// TIA Portal project "Inteligenta_szklarnia" (V15.1) (continued)
REGION Network 2: Warunki dla których okna są otwierane
   // Gdy uruchomiony jest tryb automatyczny, wartość CO2 w szklarni powinna się mieścić w zakresie nastawionego stężenia CO2 +- wartość histerezy. Okna są otwierane po spełnieniu następujących warunków: 1) gdy użytkownik załączył tryb okien na HMI, 2) gdy stężenie CO2 jest poza tym wymaganym przedziałem, 3) gdy stężenie CO2 poza szklarnią jest większe, jeśli chcemy zwiększyć ilość CO2 w szklarni oraz mniejsze, jeśli chcemy zmniejszyć ilość CO2 w szklarni, 4) gdy temperatura poza szklarnią mieści się w przedziale +-5°C temperatury nastawionej, 5) gdy wiatr wieje z prędkością nie większą niż 35km/h. Jeśli stężenie CO2 wzrośnie do niebezpiecznego poziomu 975ppm, okna również są otwierane bez względu na warunki zewnętrzne. W trybie manualnym okna otwierane są od razu po naciśnięciu przycisku do niego przypisanego.
   RUNG wire#powerrail
      Contact( #czy_automatyczny )
      I_Contact( #czy_manualny )
      wire#w1
      Contact( "HMI".System_okien_auto )
      { S7_Templates := "SrcType := Int" } LE_Contact(in1 := "Wejscia_PLC".Czujnik_wiatru, in2 := 35)
      wire#w2
      { S7_Templates := "SrcType := Int" } LT_Contact(in1 := #Histereza_plus, in2 := "HMI".Poziom_CO2_auto)
      { S7_Templates := "SrcType := Int" } GT_Contact(in1 := "Wejscia_PLC".Wewnetrzny_czujnik_CO2, in2 := "Wejscia_PLC".Zewnetrzny_czujnik_CO2)
      wire#w3
      { S7_Templates := "SrcType := Real" } InRange(min := #Zakres_temp_dol, in := "Wejscia_PLC".Temperatura_zewnetrzna, max := #Zakres_temp_gora)
      wire#w4
      I_Contact( "Siłownik_okien_zamykanie" )
      Coil( "Siłownik_okien_otwieranie" )
   END_RUNG
   RUNG wire#w2
      { S7_Templates := "SrcType := Int" } GT_Contact(in1 := #Histereza_minus, in2 := "Wejscia_PLC".Wewnetrzny_czujnik_CO2)
      { S7_Templates := "SrcType := Int" } LT_Contact(in1 := "Wejscia_PLC".Wewnetrzny_czujnik_CO2, in2 := "Wejscia_PLC".Zewnetrzny_czujnik_CO2)
   END_RUNG wire#w3
   RUNG wire#w1
      { S7_Templates := "SrcType := Int" } GE_Contact(in1 := "Wejscia_PLC".Wewnetrzny_czujnik_CO2, in2 := 975)
      { S7_Templates := "SrcType := Int" } GT_Contact(in1 := "Wejscia_PLC".Wewnetrzny_czujnik_CO2, in2 := "Wejscia_PLC".Zewnetrzny_czujnik_CO2)
   END_RUNG wire#w4
   RUNG wire#powerrail
      Contact( #czy_manualny )
      I_Contact( #czy_automatyczny )
      Contact( "HMI".Otwarcie_okien_manual )
   END_RUNG wire#w4
   // the same network as SCL:
   "Siłownik_okien_otwieranie" := ((#czy_automatyczny AND NOT #czy_manualny AND (("HMI".System_okien_auto AND ("Wejscia_PLC".Czujnik_wiatru <= 35) AND (((#Histereza_plus < "HMI".Poziom_CO2_auto) AND ("Wejscia_PLC".Wewnetrzny_czujnik_CO2 > "Wejscia_PLC".Zewnetrzny_czujnik_CO2)) OR ((#Histereza_minus > "Wejscia_PLC".Wewnetrzny_czujnik_CO2) AND ("Wejscia_PLC".Wewnetrzny_czujnik_CO2 < "Wejscia_PLC".Zewnetrzny_czujnik_CO2))) AND (#Zakres_temp_dol <= "Wejscia_PLC".Temperatura_zewnetrzna) AND ("Wejscia_PLC".Temperatura_zewnetrzna <= #Zakres_temp_gora)) OR (("Wejscia_PLC".Wewnetrzny_czujnik_CO2 >= 975) AND ("Wejscia_PLC".Wewnetrzny_czujnik_CO2 > "Wejscia_PLC".Zewnetrzny_czujnik_CO2)))) OR (#czy_manualny AND NOT #czy_automatyczny AND "HMI".Otwarcie_okien_manual)) AND NOT "Siłownik_okien_zamykanie";
END_REGION

REGION Network 3: Warunki dla których okna są zamykane
   // W trybie automatycznym okna są zamykane: 1) gdy tryb okien został wyłączony przez użytkownika, 2) gdy stężenie CO2 w szklarni wynosi zadaną wartość tego parametru +- histereza, 3) gdy stężenie CO2 poza szklarnią jest mniejsze, niż wewnątrz, jeśli chcemy zwiększyć jego ilość oraz większe, gdy chcemy zmniejszyć jego ilość, 4) gdy tempperatura zewnętrzna różni się o ponad 5°C od zadanej, 5) gdy wiatr wieje z prędkością większą niż 35km/h, 6) gdy stężenie CO2 w szklarni nie przekracza 955ppm lub przekracza, ale stężenie CO2 poza szklarnią jest większe. W trybie manualnym okna są zamykane, gdy przełączk na HMI znajdzie się w pozycji "ZAMKNIĘTE".
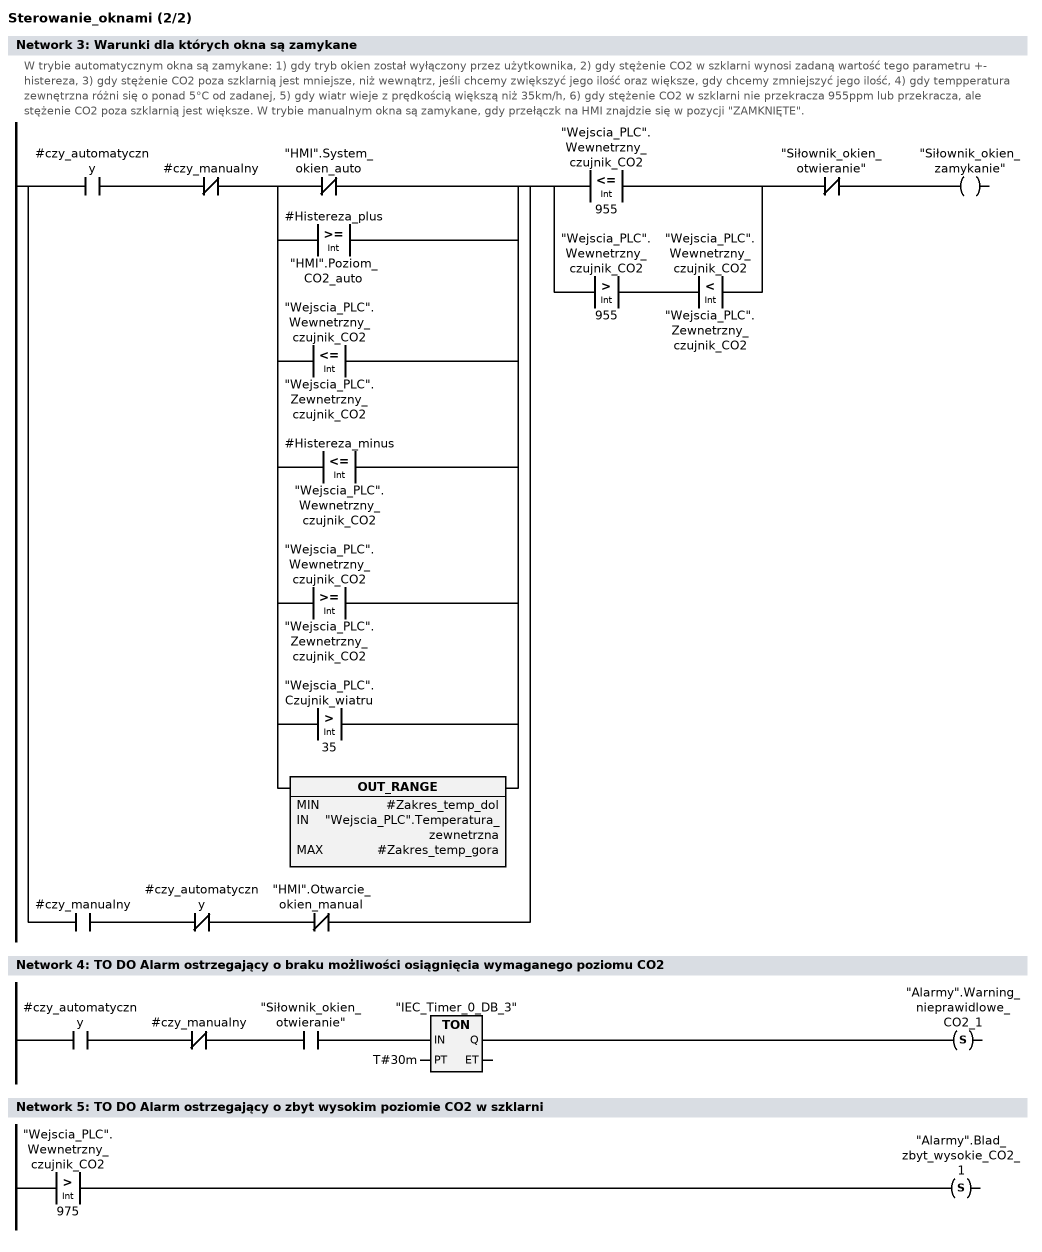
   "Siłownik_okien_zamykanie" := ((#czy_automatyczny AND NOT #czy_manualny AND (NOT "HMI".System_okien_auto OR (#Histereza_plus >= "HMI".Poziom_CO2_auto) OR ("Wejscia_PLC".Wewnetrzny_czujnik_CO2 <= "Wejscia_PLC".Zewnetrzny_czujnik_CO2) OR (#Histereza_minus <= "Wejscia_PLC".Wewnetrzny_czujnik_CO2) OR ("Wejscia_PLC".Wewnetrzny_czujnik_CO2 >= "Wejscia_PLC".Zewnetrzny_czujnik_CO2) OR ("Wejscia_PLC".Czujnik_wiatru > 35) OR ("Wejscia_PLC".Temperatura_zewnetrzna < #Zakres_temp_dol) OR ("Wejscia_PLC".Temperatura_zewnetrzna > #Zakres_temp_gora))) OR (#czy_manualny AND NOT #czy_automatyczny AND NOT "HMI".Otwarcie_okien_manual)) AND (("Wejscia_PLC".Wewnetrzny_czujnik_CO2 <= 955) OR (("Wejscia_PLC".Wewnetrzny_czujnik_CO2 > 955) AND ("Wejscia_PLC".Wewnetrzny_czujnik_CO2 < "Wejscia_PLC".Zewnetrzny_czujnik_CO2))) AND NOT "Siłownik_okien_otwieranie";
END_REGION

REGION Network 4: TO DO Alarm ostrzegający o braku możliwości osiągnięcia wymaganego poziomu CO2
   "IEC_Timer_0_DB_3".TON(IN := #czy_automatyczny AND NOT #czy_manualny AND "Siłownik_okien_otwieranie",
                          PT := T#30m);
   IF "IEC_Timer_0_DB_3".Q THEN "Alarmy".Warning_nieprawidlowe_CO2_1 := TRUE; END_IF;
END_REGION

REGION Network 5: TO DO Alarm ostrzegający o zbyt wysokim poziomie CO2 w szklarni
   RUNG wire#powerrail
      { S7_Templates := "SrcType := Int" } GT_Contact(in1 := "Wejscia_PLC".Wewnetrzny_czujnik_CO2, in2 := 975)
      S_Coil( "Alarmy".Blad_zbyt_wysokie_CO2_1 )
   END_RUNG
   // the same network as SCL:
   IF "Wejscia_PLC".Wewnetrzny_czujnik_CO2 > 975 THEN "Alarmy".Blad_zbyt_wysokie_CO2_1 := TRUE; END_IF;
END_REGION
END_FUNCTION

FUNCTION "SYMULACJA" : Void   // FC9, LAD
{ S7_Optimized_Access := 'TRUE' }
VERSION : 0.1
   VAR_INPUT
      counters : Bool;
   END_VAR
   VAR_TEMP
      temperatura_temp : Real;
      roznica_temperatur : Real;
      "wilgotność powietrza_temp" : Int;
      wilgotnosc_gleby_temp : Int;
      stezenie_CO2 : Int;
      natezenie_swiatla_temp : Int;
      odsloniecie_okna_temp : Real;
      pedkosc_wiatru_temp : Real;
      rand : Real;
      error : Bool;
      status : Int;
      sub_status : Int;
      rolety_temp : Real;
      test1 : Real;
   END_VAR
   VAR_TEMP   // added for the SCL form of the ladder/FBD networks
      _w1 : Bool;
   END_VAR
BEGIN

REGION Network 1: blok oblicza roznice temperatur
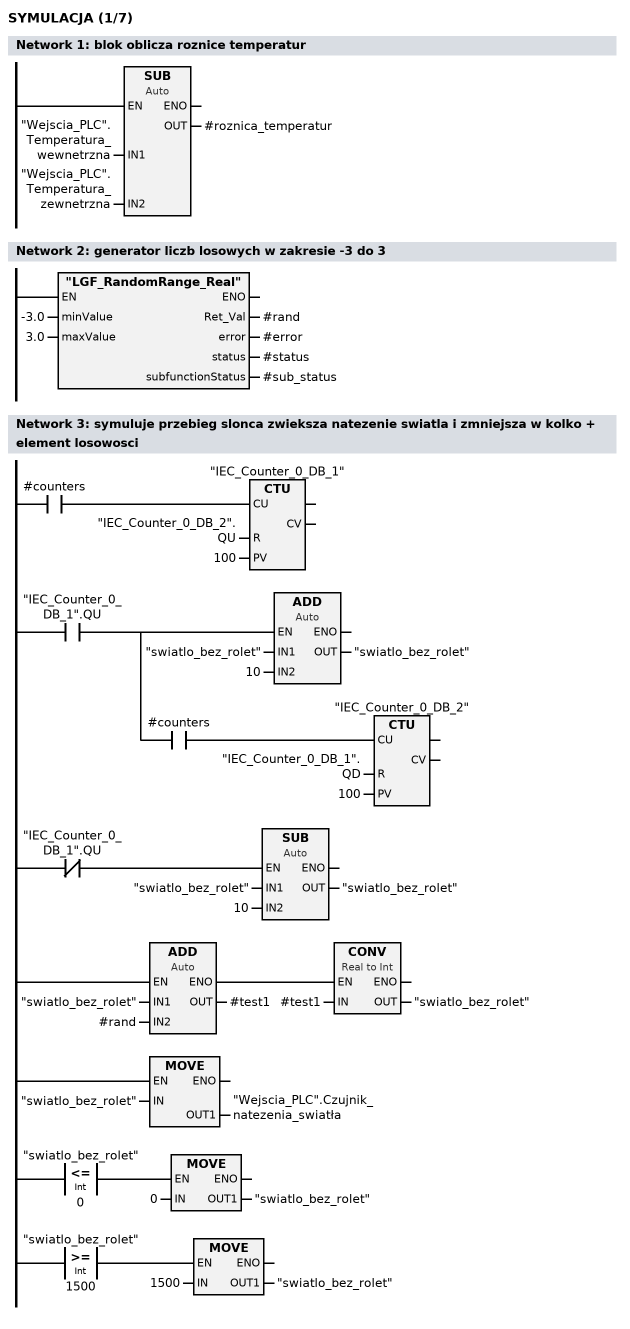
   RUNG wire#powerrail
      { S7_GenerateENO := "TRUE" } Sub(in1 := "Wejscia_PLC".Temperatura_wewnetrzna, in2 := "Wejscia_PLC".Temperatura_zewnetrzna, out => #roznica_temperatur)
   END_RUNG
   // the same network as SCL:
   #roznica_temperatur := "Wejscia_PLC".Temperatura_wewnetrzna - "Wejscia_PLC".Temperatura_zewnetrzna;
END_REGION

REGION Network 2: generator liczb losowych w zakresie -3 do 3
   RUNG wire#powerrail
      "LGF_RandomRange_Real"(minValue := -3.0, maxValue := 3.0, Ret_Val => #rand, error => #error, status => #status, subfunctionStatus => #sub_status)
   END_RUNG
   // the same network as SCL:
   #rand := "LGF_RandomRange_Real"(minValue := -3.0,
                           maxValue := 3.0,
                           error => #error,
                           status => #status,
                           subfunctionStatus => #sub_status);
END_REGION

REGION Network 3: symuluje przebieg slonca zwieksza natezenie swiatla i zmniejsza w kolko + element losowosci
   // ENO of a box is taken as its EN; it also drops when the box reports an error
   "IEC_Counter_0_DB_1".CTU(CU := #counters, R := "IEC_Counter_0_DB_2".QU, PV := 100);
   IF "IEC_Counter_0_DB_1".QU THEN "swiatlo_bez_rolet" := "swiatlo_bez_rolet" + 10; END_IF;
   "IEC_Counter_0_DB_2".CTU(CU := "IEC_Counter_0_DB_1".QU AND #counters,
                           R := "IEC_Counter_0_DB_1".QD,
                           PV := 100);
   IF NOT "IEC_Counter_0_DB_1".QU THEN "swiatlo_bez_rolet" := "swiatlo_bez_rolet" - 10; END_IF;
   #test1 := "swiatlo_bez_rolet" + #rand;
   "swiatlo_bez_rolet" := REAL_TO_INT(#test1);
   "Wejscia_PLC".Czujnik_natezenia_swiatła := "swiatlo_bez_rolet";
   IF "swiatlo_bez_rolet" <= 0 THEN "swiatlo_bez_rolet" := 0; END_IF;
   IF "swiatlo_bez_rolet" >= 1500 THEN "swiatlo_bez_rolet" := 1500; END_IF;
END_REGION

REGION Network 4: funkcja oblicza liniową zależność natężenia światła od zasłonięcia rolet
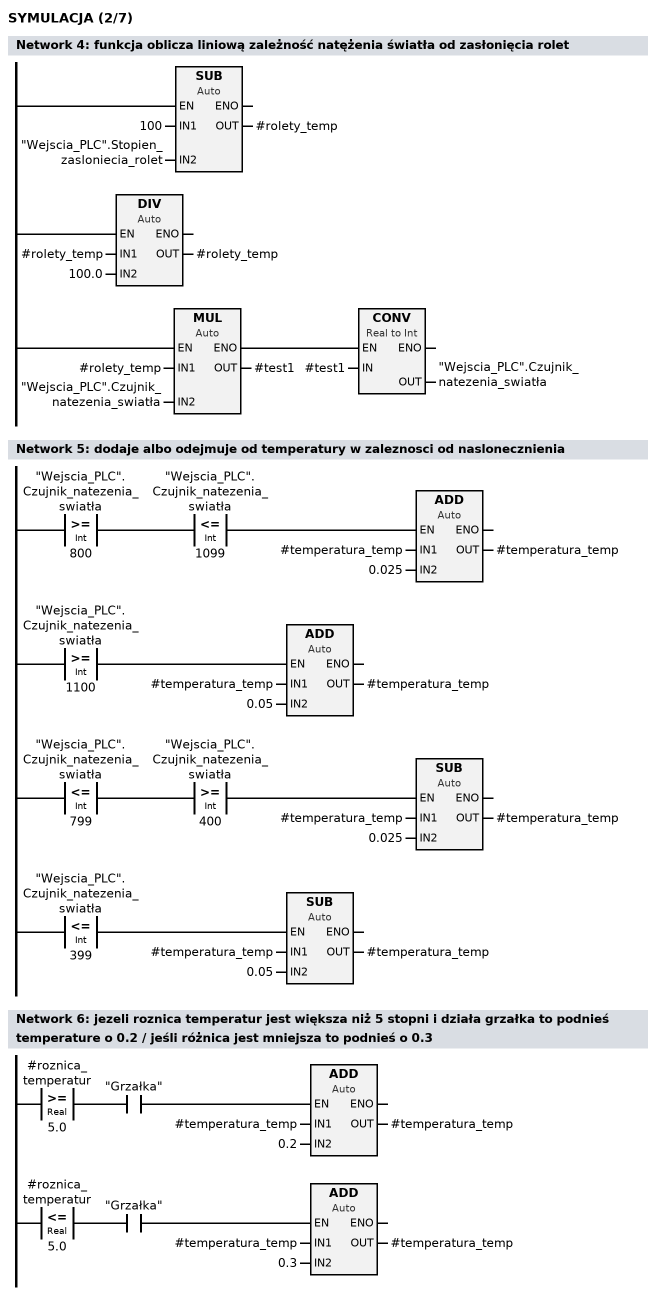
   RUNG wire#powerrail
      { S7_GenerateENO := "TRUE" } Sub(in1 := 100, in2 := "Wejscia_PLC".Stopien_zasloniecia_rolet, out => #rolety_temp)
   END_RUNG
   RUNG wire#powerrail
      { S7_GenerateENO := "TRUE" } Div(in1 := #rolety_temp, in2 := 100.0, out => #rolety_temp)
   END_RUNG
   RUNG wire#powerrail
      { S7_GenerateENO := "TRUE" } Mul(in1 := #rolety_temp, in2 := "Wejscia_PLC".Czujnik_natezenia_swiatła, out => #test1)
      { S7_Templates := "[SrcType := Real, DestType := Int]"; S7_GenerateENO := "TRUE" } Convert(in := #test1, out => "Wejscia_PLC".Czujnik_natezenia_swiatła)
   END_RUNG
   // the same network as SCL:
   // ENO of a box is taken as its EN; it also drops when the box reports an error
   #rolety_temp := 100 - "Wejscia_PLC".Stopien_zasloniecia_rolet;
   #rolety_temp := #rolety_temp / 100.0;
   #test1 := #rolety_temp * "Wejscia_PLC".Czujnik_natezenia_swiatła;
   "Wejscia_PLC".Czujnik_natezenia_swiatła := REAL_TO_INT(#test1);
END_REGION

REGION Network 5: dodaje albo odejmuje od temperatury w zaleznosci od naslonecznienia
   RUNG wire#powerrail
      { S7_Templates := "SrcType := Int" } GE_Contact(in1 := "Wejscia_PLC".Czujnik_natezenia_swiatła, in2 := 800)
      { S7_Templates := "SrcType := Int" } LE_Contact(in1 := "Wejscia_PLC".Czujnik_natezenia_swiatła, in2 := 1099)
      { S7_GenerateENO := "TRUE" } Add(in1 := #temperatura_temp, in2 := 0.025, out => #temperatura_temp)
   END_RUNG
   RUNG wire#powerrail
      { S7_Templates := "SrcType := Int" } GE_Contact(in1 := "Wejscia_PLC".Czujnik_natezenia_swiatła, in2 := 1100)
      { S7_GenerateENO := "TRUE" } Add(in1 := #temperatura_temp, in2 := 0.05, out => #temperatura_temp)
   END_RUNG
   RUNG wire#powerrail
      { S7_Templates := "SrcType := Int" } LE_Contact(in1 := "Wejscia_PLC".Czujnik_natezenia_swiatła, in2 := 799)
      { S7_Templates := "SrcType := Int" } GE_Contact(in1 := "Wejscia_PLC".Czujnik_natezenia_swiatła, in2 := 400)
      { S7_GenerateENO := "TRUE" } Sub(in1 := #temperatura_temp, in2 := 0.025, out => #temperatura_temp)
   END_RUNG
   RUNG wire#powerrail
      { S7_Templates := "SrcType := Int" } LE_Contact(in1 := "Wejscia_PLC".Czujnik_natezenia_swiatła, in2 := 399)
      { S7_GenerateENO := "TRUE" } Sub(in1 := #temperatura_temp, in2 := 0.05, out => #temperatura_temp)
   END_RUNG
   // the same network as SCL:
   IF ("Wejscia_PLC".Czujnik_natezenia_swiatła >= 800) AND ("Wejscia_PLC".Czujnik_natezenia_swiatła <= 1099) THEN
       #temperatura_temp := #temperatura_temp + 0.025;
   END_IF;
   IF "Wejscia_PLC".Czujnik_natezenia_swiatła >= 1100 THEN
       #temperatura_temp := #temperatura_temp + 0.05;
   END_IF;
   IF ("Wejscia_PLC".Czujnik_natezenia_swiatła <= 799) AND ("Wejscia_PLC".Czujnik_natezenia_swiatła >= 400) THEN
       #temperatura_temp := #temperatura_temp - 0.025;
   END_IF;
   IF "Wejscia_PLC".Czujnik_natezenia_swiatła <= 399 THEN
       #temperatura_temp := #temperatura_temp - 0.05;
   END_IF;
END_REGION

REGION Network 6: jezeli roznica temperatur jest większa niż 5 stopni i działa grzałka to podnieś temperature o 0.2 / jeśli różnica jest mniejsza to podnieś o 0.3
   RUNG wire#powerrail
      { S7_Templates := "SrcType := Real" } GE_Contact(in1 := #roznica_temperatur, in2 := 5.0)
      Contact( "Grzałka" )
      { S7_GenerateENO := "TRUE" } Add(in1 := #temperatura_temp, in2 := 0.2, out => #temperatura_temp)
   END_RUNG
   RUNG wire#powerrail
      { S7_Templates := "SrcType := Real" } LE_Contact(in1 := #roznica_temperatur, in2 := 5.0)
      Contact( "Grzałka" )
      { S7_GenerateENO := "TRUE" } Add(in1 := #temperatura_temp, in2 := 0.3, out => #temperatura_temp)
   END_RUNG
   // the same network as SCL:
   IF (#roznica_temperatur >= 5.0) AND "Grzałka" THEN #temperatura_temp := #temperatura_temp + 0.2; END_IF;
   IF (#roznica_temperatur <= 5.0) AND "Grzałka" THEN #temperatura_temp := #temperatura_temp + 0.3; END_IF;
END_REGION

REGION Network 7: jezeli działa wentylator to obniż temperature o 0.1
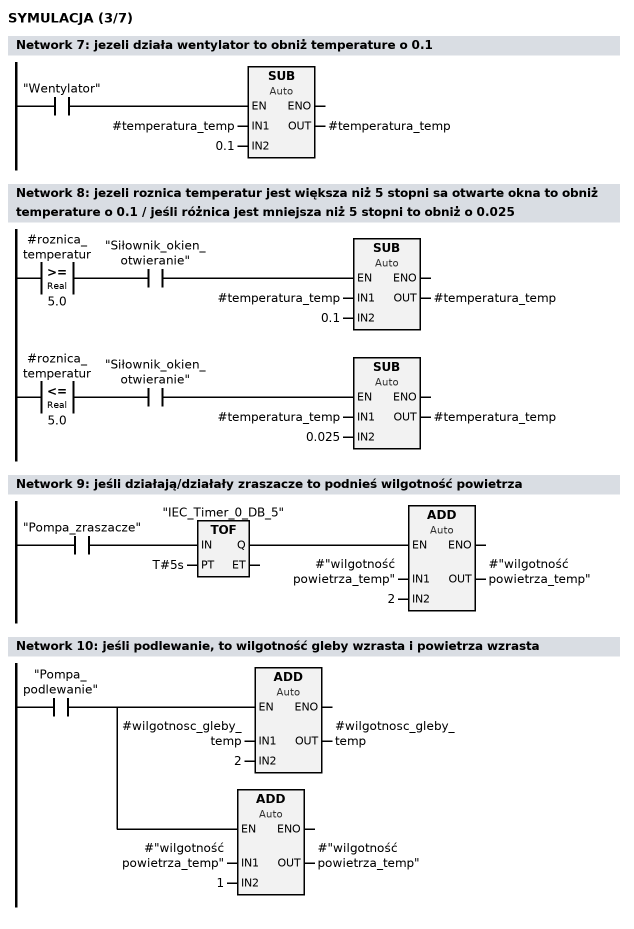
   RUNG wire#powerrail
      Contact( "Wentylator" )
      { S7_GenerateENO := "TRUE" } Sub(in1 := #temperatura_temp, in2 := 0.1, out => #temperatura_temp)
   END_RUNG
   // the same network as SCL:
   IF "Wentylator" THEN #temperatura_temp := #temperatura_temp - 0.1; END_IF;
END_REGION

REGION Network 8: jezeli roznica temperatur jest większa niż 5 stopni sa otwarte okna to obniż temperature o 0.1 / jeśli różnica jest mniejsza niż 5 stopni to obniż o 0.025
   RUNG wire#powerrail
      { S7_Templates := "SrcType := Real" } GE_Contact(in1 := #roznica_temperatur, in2 := 5.0)
      Contact( "Siłownik_okien_otwieranie" )
      { S7_GenerateENO := "TRUE" } Sub(in1 := #temperatura_temp, in2 := 0.1, out => #temperatura_temp)
   END_RUNG
   RUNG wire#powerrail
      { S7_Templates := "SrcType := Real" } LE_Contact(in1 := #roznica_temperatur, in2 := 5.0)
      Contact( "Siłownik_okien_otwieranie" )
      { S7_GenerateENO := "TRUE" } Sub(in1 := #temperatura_temp, in2 := 0.025, out => #temperatura_temp)
   END_RUNG
   // the same network as SCL:
   IF (#roznica_temperatur >= 5.0) AND "Siłownik_okien_otwieranie" THEN
       #temperatura_temp := #temperatura_temp - 0.1;
   END_IF;
   IF (#roznica_temperatur <= 5.0) AND "Siłownik_okien_otwieranie" THEN
       #temperatura_temp := #temperatura_temp - 0.025;
   END_IF;
END_REGION

REGION Network 9: jeśli działają/działały zraszacze to podnieś wilgotność powietrza
   "IEC_Timer_0_DB_5".TOF(IN := "Pompa_zraszacze", PT := T#5s);
   IF "IEC_Timer_0_DB_5".Q THEN #"wilgotność powietrza_temp" := #"wilgotność powietrza_temp" + 2; END_IF;
END_REGION

REGION Network 10: jeśli podlewanie, to wilgotność gleby wzrasta i powietrza wzrasta
   RUNG wire#powerrail
      Contact( "Pompa_podlewanie" )
      wire#w1
      { S7_GenerateENO := "TRUE" } Add(in1 := #wilgotnosc_gleby_temp, in2 := 2, out => #wilgotnosc_gleby_temp)
   END_RUNG
   RUNG wire#w1
      { S7_GenerateENO := "TRUE" } Add(in1 := #"wilgotność powietrza_temp", in2 := 1, out => #"wilgotność powietrza_temp")
   END_RUNG
   // the same network as SCL:
   IF "Pompa_podlewanie" THEN
       #wilgotnosc_gleby_temp := #wilgotnosc_gleby_temp + 2;
       #"wilgotność powietrza_temp" := #"wilgotność powietrza_temp" + 1;
   END_IF;
END_REGION

REGION Network 11: realizacja zaleznosci odslaniania i zaslaniania rolet, od stopnia zasłonięcia
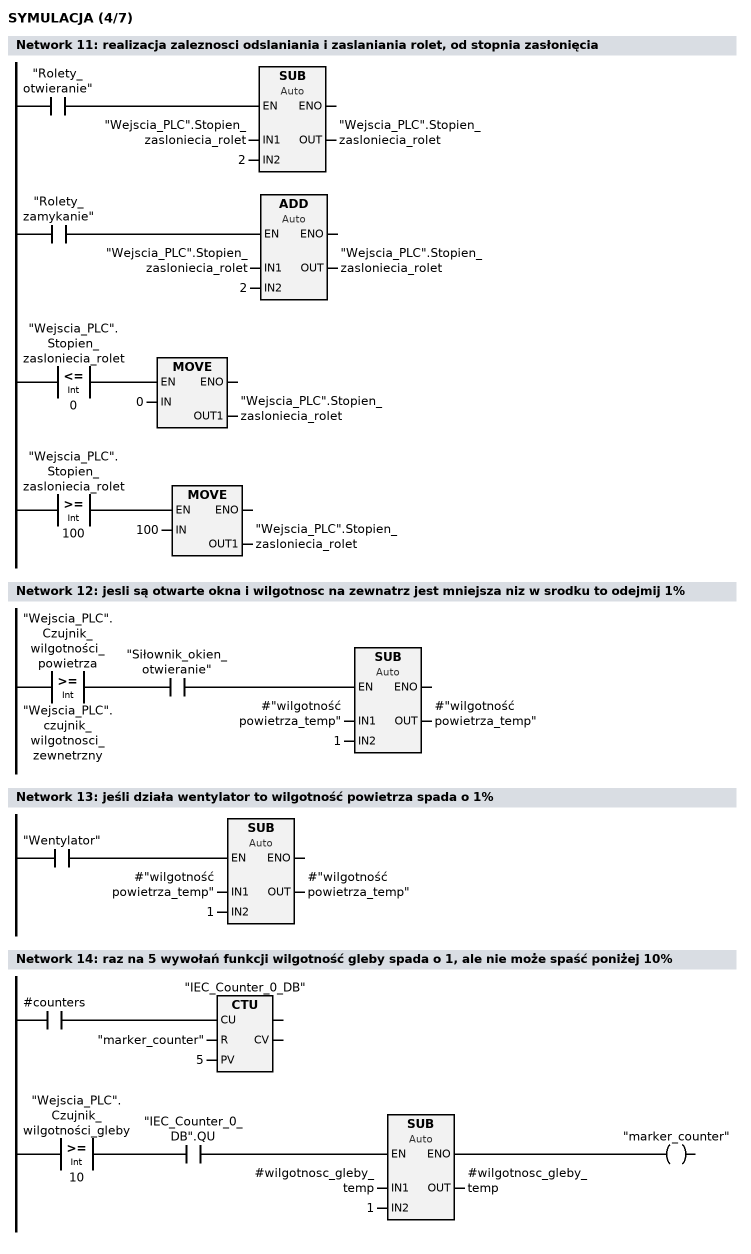
   RUNG wire#powerrail
      Contact( "Rolety_otwieranie" )
      { S7_GenerateENO := "TRUE" } Sub(in1 := "Wejscia_PLC".Stopien_zasloniecia_rolet, in2 := 2, out => "Wejscia_PLC".Stopien_zasloniecia_rolet)
   END_RUNG
   RUNG wire#powerrail
      Contact( "Rolety_zamykanie" )
      { S7_GenerateENO := "TRUE" } Add(in1 := "Wejscia_PLC".Stopien_zasloniecia_rolet, in2 := 2, out => "Wejscia_PLC".Stopien_zasloniecia_rolet)
   END_RUNG
   RUNG wire#powerrail
      { S7_Templates := "SrcType := Int" } LE_Contact(in1 := "Wejscia_PLC".Stopien_zasloniecia_rolet, in2 := 0)
      { S7_GenerateENO := "TRUE" } Move(in := 0, out1 => "Wejscia_PLC".Stopien_zasloniecia_rolet)
   END_RUNG
   RUNG wire#powerrail
      { S7_Templates := "SrcType := Int" } GE_Contact(in1 := "Wejscia_PLC".Stopien_zasloniecia_rolet, in2 := 100)
      { S7_GenerateENO := "TRUE" } Move(in := 100, out1 => "Wejscia_PLC".Stopien_zasloniecia_rolet)
   END_RUNG
   // the same network as SCL:
   IF "Rolety_otwieranie" THEN
       "Wejscia_PLC".Stopien_zasloniecia_rolet := "Wejscia_PLC".Stopien_zasloniecia_rolet - 2;
   END_IF;
   IF "Rolety_zamykanie" THEN
       "Wejscia_PLC".Stopien_zasloniecia_rolet := "Wejscia_PLC".Stopien_zasloniecia_rolet + 2;
   END_IF;
   IF "Wejscia_PLC".Stopien_zasloniecia_rolet <= 0 THEN "Wejscia_PLC".Stopien_zasloniecia_rolet := 0; END_IF;
   IF "Wejscia_PLC".Stopien_zasloniecia_rolet >= 100 THEN
       "Wejscia_PLC".Stopien_zasloniecia_rolet := 100;
   END_IF;
END_REGION

REGION Network 12: jesli są otwarte okna i wilgotnosc na zewnatrz jest mniejsza niz w srodku to odejmij 1%
   RUNG wire#powerrail
      { S7_Templates := "SrcType := Int" } GE_Contact(in1 := "Wejscia_PLC".Czujnik_wilgotności_powietrza, in2 := "Wejscia_PLC".czujnik_wilgotnosci_zewnetrzny)
      Contact( "Siłownik_okien_otwieranie" )
      { S7_GenerateENO := "TRUE" } Sub(in1 := #"wilgotność powietrza_temp", in2 := 1, out => #"wilgotność powietrza_temp")
   END_RUNG
   // the same network as SCL:
   IF ("Wejscia_PLC".Czujnik_wilgotności_powietrza >= "Wejscia_PLC".czujnik_wilgotnosci_zewnetrzny) AND "Siłownik_okien_otwieranie" THEN
       #"wilgotność powietrza_temp" := #"wilgotność powietrza_temp" - 1;
   END_IF;
END_REGION

REGION Network 13: jeśli działa wentylator to wilgotność powietrza spada o 1%
   RUNG wire#powerrail
      Contact( "Wentylator" )
      { S7_GenerateENO := "TRUE" } Sub(in1 := #"wilgotność powietrza_temp", in2 := 1, out => #"wilgotność powietrza_temp")
   END_RUNG
   // the same network as SCL:
   IF "Wentylator" THEN #"wilgotność powietrza_temp" := #"wilgotność powietrza_temp" - 1; END_IF;
END_REGION

REGION Network 14: raz na 5 wywołań funkcji wilgotność gleby spada o 1, ale nie może spaść poniżej 10%
   // ENO of a box is taken as its EN; it also drops when the box reports an error
   "IEC_Counter_0_DB".CTU(CU := #counters, R := "marker_counter", PV := 5);
   #_w1 := ("Wejscia_PLC".Czujnik_wilgotności_gleby >= 10) AND "IEC_Counter_0_DB".QU;
   IF #_w1 THEN #wilgotnosc_gleby_temp := #wilgotnosc_gleby_temp - 1; END_IF;
   "marker_counter" := #_w1;
END_REGION

REGION Network 15: jeśli stężenie na zewnątrz jest mniejsze, a są otwarte okna to zmniejsz stężenie CO2
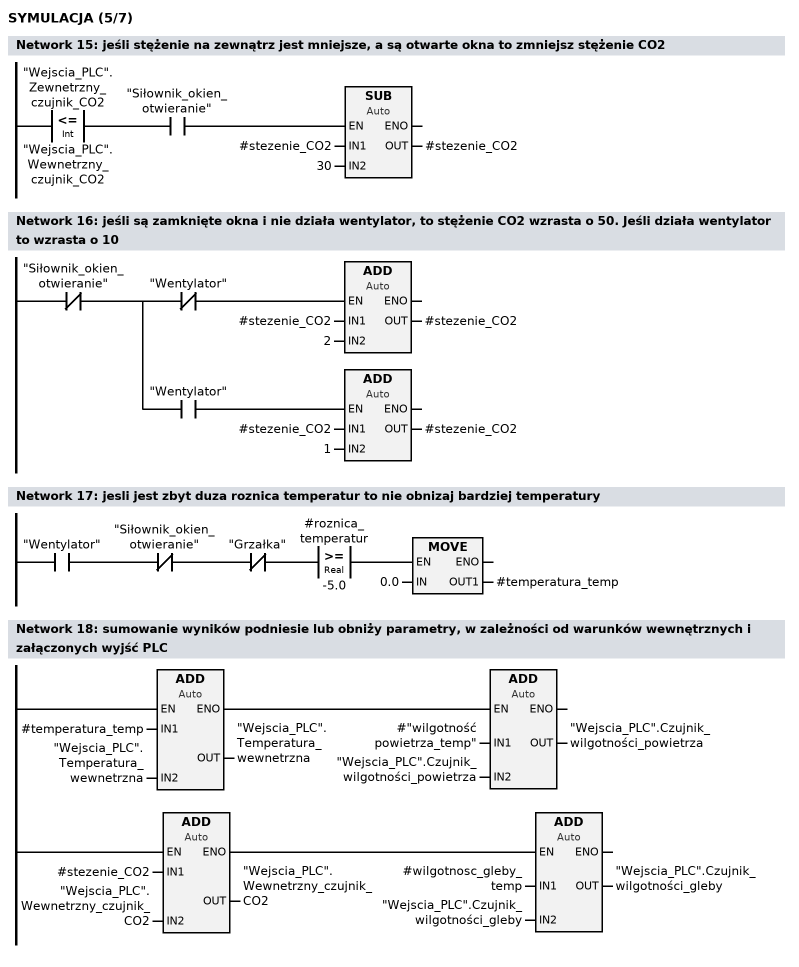
   RUNG wire#powerrail
      { S7_Templates := "SrcType := Int" } LE_Contact(in1 := "Wejscia_PLC".Zewnetrzny_czujnik_CO2, in2 := "Wejscia_PLC".Wewnetrzny_czujnik_CO2)
      Contact( "Siłownik_okien_otwieranie" )
      { S7_GenerateENO := "TRUE" } Sub(in1 := #stezenie_CO2, in2 := 30, out => #stezenie_CO2)
   END_RUNG
   // the same network as SCL:
   IF ("Wejscia_PLC".Zewnetrzny_czujnik_CO2 <= "Wejscia_PLC".Wewnetrzny_czujnik_CO2) AND "Siłownik_okien_otwieranie" THEN
       #stezenie_CO2 := #stezenie_CO2 - 30;
   END_IF;
END_REGION

REGION Network 16: jeśli są zamknięte okna i nie działa wentylator, to stężenie CO2 wzrasta o 50. Jeśli działa wentylator to wzrasta o 10
   RUNG wire#powerrail
      I_Contact( "Siłownik_okien_otwieranie" )
      wire#w1
      I_Contact( "Wentylator" )
      { S7_GenerateENO := "TRUE" } Add(in1 := #stezenie_CO2, in2 := 2, out => #stezenie_CO2)
   END_RUNG
   RUNG wire#w1
      Contact( "Wentylator" )
      { S7_GenerateENO := "TRUE" } Add(in1 := #stezenie_CO2, in2 := 1, out => #stezenie_CO2)
   END_RUNG
   // the same network as SCL:
   #_w1 := NOT "Siłownik_okien_otwieranie";
   IF #_w1 AND NOT "Wentylator" THEN #stezenie_CO2 := #stezenie_CO2 + 2; END_IF;
   IF #_w1 AND "Wentylator" THEN #stezenie_CO2 := #stezenie_CO2 + 1; END_IF;
END_REGION

REGION Network 17: jesli jest zbyt duza roznica temperatur to nie obnizaj bardziej temperatury
   RUNG wire#powerrail
      Contact( "Wentylator" )
      I_Contact( "Siłownik_okien_otwieranie" )
      I_Contact( "Grzałka" )
      { S7_Templates := "SrcType := Real" } GE_Contact(in1 := #roznica_temperatur, in2 := -5.0)
      { S7_GenerateENO := "TRUE" } Move(in := 0.0, out1 => #temperatura_temp)
   END_RUNG
   // the same network as SCL:
   IF "Wentylator" AND NOT "Siłownik_okien_otwieranie" AND NOT "Grzałka" AND (#roznica_temperatur >= (-5.0)) THEN
       #temperatura_temp := 0.0;
   END_IF;
END_REGION

REGION Network 18: sumowanie wyników podniesie lub obniży parametry, w zależności od warunków wewnętrznych i załączonych wyjść PLC
   RUNG wire#powerrail
      { S7_GenerateENO := "TRUE" } Add(in1 := #temperatura_temp, in2 := "Wejscia_PLC".Temperatura_wewnetrzna, out => "Wejscia_PLC".Temperatura_wewnetrzna)
      { S7_GenerateENO := "TRUE" } Add(in1 := #"wilgotność powietrza_temp", in2 := "Wejscia_PLC".Czujnik_wilgotności_powietrza, out => "Wejscia_PLC".Czujnik_wilgotności_powietrza)
   END_RUNG
   RUNG wire#powerrail
      { S7_GenerateENO := "TRUE" } Add(in1 := #stezenie_CO2, in2 := "Wejscia_PLC".Wewnetrzny_czujnik_CO2, out => "Wejscia_PLC".Wewnetrzny_czujnik_CO2)
      { S7_GenerateENO := "TRUE" } Add(in1 := #wilgotnosc_gleby_temp, in2 := "Wejscia_PLC".Czujnik_wilgotności_gleby, out => "Wejscia_PLC".Czujnik_wilgotności_gleby)
   END_RUNG
   // the same network as SCL:
   // ENO of a box is taken as its EN; it also drops when the box reports an error
   "Wejscia_PLC".Temperatura_wewnetrzna := #temperatura_temp + "Wejscia_PLC".Temperatura_wewnetrzna;
   "Wejscia_PLC".Czujnik_wilgotności_powietrza := #"wilgotność powietrza_temp" + "Wejscia_PLC".Czujnik_wilgotności_powietrza;
   "Wejscia_PLC".Wewnetrzny_czujnik_CO2 := #stezenie_CO2 + "Wejscia_PLC".Wewnetrzny_czujnik_CO2;
   "Wejscia_PLC".Czujnik_wilgotności_gleby := #wilgotnosc_gleby_temp + "Wejscia_PLC".Czujnik_wilgotności_gleby;
END_REGION

REGION Network 19: zabezpieczenie, przed przekroczeniem wartości krytycznych czujników + zabezpieczenia fizyczne np. procenty tylko w zakresie(0-100)
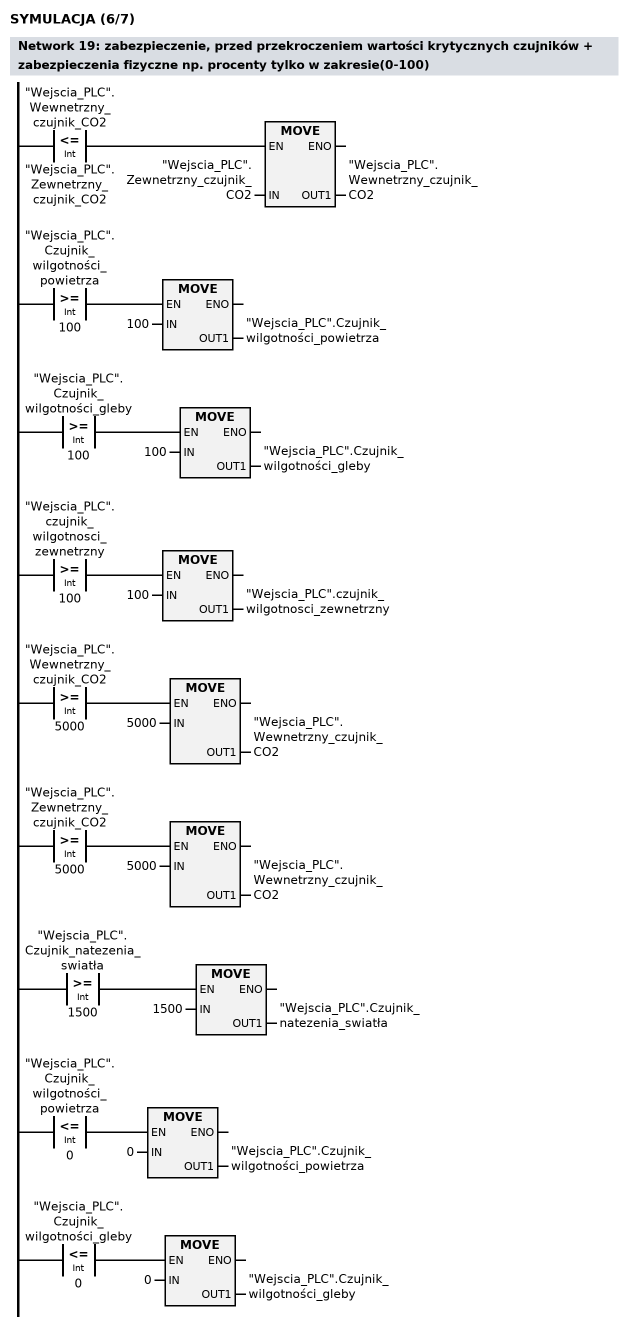
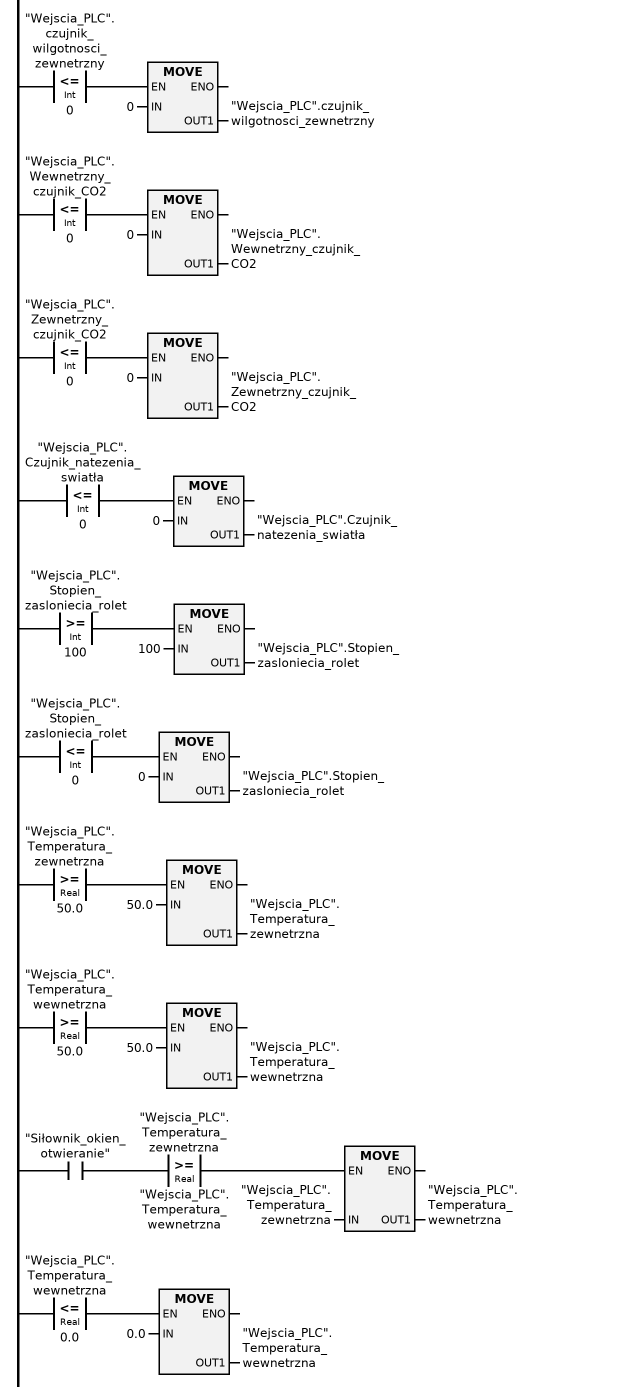
   RUNG wire#powerrail
      { S7_Templates := "SrcType := Int" } LE_Contact(in1 := "Wejscia_PLC".Wewnetrzny_czujnik_CO2, in2 := "Wejscia_PLC".Zewnetrzny_czujnik_CO2)
      { S7_GenerateENO := "TRUE" } Move(in := "Wejscia_PLC".Zewnetrzny_czujnik_CO2, out1 => "Wejscia_PLC".Wewnetrzny_czujnik_CO2)
   END_RUNG
   RUNG wire#powerrail
      { S7_Templates := "SrcType := Int" } GE_Contact(in1 := "Wejscia_PLC".Czujnik_wilgotności_powietrza, in2 := 100)
      { S7_GenerateENO := "TRUE" } Move(in := 100, out1 => "Wejscia_PLC".Czujnik_wilgotności_powietrza)
   END_RUNG
   RUNG wire#powerrail
      { S7_Templates := "SrcType := Int" } GE_Contact(in1 := "Wejscia_PLC".Czujnik_wilgotności_gleby, in2 := 100)
      { S7_GenerateENO := "TRUE" } Move(in := 100, out1 => "Wejscia_PLC".Czujnik_wilgotności_gleby)
   END_RUNG
   RUNG wire#powerrail
      { S7_Templates := "SrcType := Int" } GE_Contact(in1 := "Wejscia_PLC".czujnik_wilgotnosci_zewnetrzny, in2 := 100)
      { S7_GenerateENO := "TRUE" } Move(in := 100, out1 => "Wejscia_PLC".czujnik_wilgotnosci_zewnetrzny)
   END_RUNG
   RUNG wire#powerrail
      { S7_Templates := "SrcType := Int" } GE_Contact(in1 := "Wejscia_PLC".Wewnetrzny_czujnik_CO2, in2 := 5000)
      { S7_GenerateENO := "TRUE" } Move(in := 5000, out1 => "Wejscia_PLC".Wewnetrzny_czujnik_CO2)
   END_RUNG
   RUNG wire#powerrail
      { S7_Templates := "SrcType := Int" } GE_Contact(in1 := "Wejscia_PLC".Zewnetrzny_czujnik_CO2, in2 := 5000)
      { S7_GenerateENO := "TRUE" } Move(in := 5000, out1 => "Wejscia_PLC".Wewnetrzny_czujnik_CO2)
   END_RUNG
   RUNG wire#powerrail
      { S7_Templates := "SrcType := Int" } GE_Contact(in1 := "Wejscia_PLC".Czujnik_natezenia_swiatła, in2 := 1500)
      { S7_GenerateENO := "TRUE" } Move(in := 1500, out1 => "Wejscia_PLC".Czujnik_natezenia_swiatła)
   END_RUNG
   RUNG wire#powerrail
      { S7_Templates := "SrcType := Int" } LE_Contact(in1 := "Wejscia_PLC".Czujnik_wilgotności_powietrza, in2 := 0)
      { S7_GenerateENO := "TRUE" } Move(in := 0, out1 => "Wejscia_PLC".Czujnik_wilgotności_powietrza)
   END_RUNG
   RUNG wire#powerrail
      { S7_Templates := "SrcType := Int" } LE_Contact(in1 := "Wejscia_PLC".Czujnik_wilgotności_gleby, in2 := 0)
      { S7_GenerateENO := "TRUE" } Move(in := 0, out1 => "Wejscia_PLC".Czujnik_wilgotności_gleby)
   END_RUNG
   RUNG wire#powerrail
      { S7_Templates := "SrcType := Int" } LE_Contact(in1 := "Wejscia_PLC".czujnik_wilgotnosci_zewnetrzny, in2 := 0)
      { S7_GenerateENO := "TRUE" } Move(in := 0, out1 => "Wejscia_PLC".czujnik_wilgotnosci_zewnetrzny)
   END_RUNG
   RUNG wire#powerrail
      { S7_Templates := "SrcType := Int" } LE_Contact(in1 := "Wejscia_PLC".Wewnetrzny_czujnik_CO2, in2 := 0)
      { S7_GenerateENO := "TRUE" } Move(in := 0, out1 => "Wejscia_PLC".Wewnetrzny_czujnik_CO2)
   END_RUNG
   RUNG wire#powerrail
      { S7_Templates := "SrcType := Int" } LE_Contact(in1 := "Wejscia_PLC".Zewnetrzny_czujnik_CO2, in2 := 0)
      { S7_GenerateENO := "TRUE" } Move(in := 0, out1 => "Wejscia_PLC".Zewnetrzny_czujnik_CO2)
   END_RUNG
   RUNG wire#powerrail
      { S7_Templates := "SrcType := Int" } LE_Contact(in1 := "Wejscia_PLC".Czujnik_natezenia_swiatła, in2 := 0)
      { S7_GenerateENO := "TRUE" } Move(in := 0, out1 => "Wejscia_PLC".Czujnik_natezenia_swiatła)
   END_RUNG
   RUNG wire#powerrail
      { S7_Templates := "SrcType := Int" } GE_Contact(in1 := "Wejscia_PLC".Stopien_zasloniecia_rolet, in2 := 100)
      { S7_GenerateENO := "TRUE" } Move(in := 100, out1 => "Wejscia_PLC".Stopien_zasloniecia_rolet)
   END_RUNG
   RUNG wire#powerrail
      { S7_Templates := "SrcType := Int" } LE_Contact(in1 := "Wejscia_PLC".Stopien_zasloniecia_rolet, in2 := 0)
      { S7_GenerateENO := "TRUE" } Move(in := 0, out1 => "Wejscia_PLC".Stopien_zasloniecia_rolet)
   END_RUNG
   RUNG wire#powerrail
      { S7_Templates := "SrcType := Real" } GE_Contact(in1 := "Wejscia_PLC".Temperatura_zewnetrzna, in2 := 50.0)
      { S7_GenerateENO := "TRUE" } Move(in := 50.0, out1 => "Wejscia_PLC".Temperatura_zewnetrzna)
   END_RUNG
   RUNG wire#powerrail
      { S7_Templates := "SrcType := Real" } GE_Contact(in1 := "Wejscia_PLC".Temperatura_wewnetrzna, in2 := 50.0)
      { S7_GenerateENO := "TRUE" } Move(in := 50.0, out1 => "Wejscia_PLC".Temperatura_wewnetrzna)
   END_RUNG